
screen "手动设置" 1280x733, template "模板_1"
   on GenerateScreen: SetTag("变量_100", 8)
   Button "HmiScreenItemData_1" at 1116,125 size 159x47; TextOn '向后 / 後向き / 뒤로'; TextOff '向后 / 後向き / 뒤로'
      on Release: ActivateScreen("手动画面", 0)
   IOField "IO 域_20" at 80,185 size 120x41; FormatPattern 99999999
      on Activate: function_f41c6f6c("变量_1")
      ProcessValue <- "ST_HMI_Var_HMI_r64Velocity_Jog_Chuche"
   TextField "文本域_19" at 848,56 size 245x25; Text '当前登录用户 / 目前ログオン中のユーザー / 현재 로그인 사용자'
   IOField "IO 域_15" at 914,98 size 122x41; FormatPattern ?????????????
      ProcessValue <- "user_name"
   IOField "IO 域_2" at 80,417 size 120x41; FormatPattern 99999999
      ProcessValue <- "ST_HMI_Var_HMI_r64Velocity_Jog_JinChe"
   IOField "IO 域_3" at 232,417 size 120x41; FormatPattern 999999999
      ProcessValue <- "ST_HMI_Var_HMI_r64Velocity_Jog_JiaNian"
   IOField "IO 域_5" at 384,417 size 120x41; FormatPattern 999999999
      ProcessValue <- "ST_HMI_Var_HMI_r64Velocity_Jog_JuanRao"
   IOField "IO 域_4" at 232,185 size 120x41; FormatPattern 99999999
      ProcessValue <- "ST_HMI_Var_HMI_r64Velocity_Jog_SongTiao"
   IOField "IO 域_16" at 384,185 size 120x41; FormatPattern 999999999
      ProcessValue <- "ST_HMI_Var_HMI_r64Velocity_Jog_TuiRao"
   IOField "IO 域_6" at 536,416 size 120x41; Authorization "User administration"; FormatPattern 99999999
      ProcessValue <- "ST_HMI_Var_HMI_r64Velocity_Jog_ChengXing_Up"
   IOField "IO 域_7" at 536,186 size 120x41; Authorization "User administration"; FormatPattern 99999999
      ProcessValue <- "ST_HMI_Var_HMI_r64Velocity_Jog_ChengXing_Down"
   IOField "IO 域_9" at 688,184 size 120x41; Authorization "User administration"; FormatPattern 99999999
      ProcessValue <- "ST_HMI_Var_HMI_r64Velocity_Jog_ZhangLi_Up"
   IOField "IO 域_10" at 688,416 size 120x41; Authorization "User administration"; FormatPattern 99999999
      ProcessValue <- "ST_HMI_Var_HMI_r64Velocity_Jog_ZhangLi_Down"
   IOField "IO 域_21" at 80,253 size 120x41; FormatPattern 99999999
      on Activate: function_f41c6f6c("变量_1")
      ProcessValue <- "ST_HMI_Var_HMI_r64AccVelocity_Jog_ChuChe"
   IOField "IO 域_8" at 80,485 size 120x41; FormatPattern 99999999
      ProcessValue <- "ST_HMI_Var_HMI_r64AccVelocity_Jog_JinChe"
   Button "OBJECT_119" at 328,588 size 177x68; TextOff '选择市电模式 / EXIT / 買電モードの選択 / 일반전력'; Authorization "Operate_5"
      on Press: SetBit("ST_HMI_Var_HMI_Bo_Feed_On_Off_Select")
      Appearance <- "ST_HMI_Var_HMI_Bo_Feed_On_Off_Select"
   Button "OBJECT_120" at 573,588 size 177x68; TextOff '选择发电模式 / EXIT / 発電モードの選択 / 발전기 전력'; Authorization "Operate_5"
      on Press: ResetBit("ST_HMI_Var_HMI_Bo_Feed_On_Off_Select")
      Appearance <- "ST_HMI_Var_HMI_Bo_Feed_On_Off_Select"
   Button "OBJECT_5" at 80,80 size 120x80; TextOff '出车 / EXIT / 出機 / 외진'
      on Release: ResetBit("ST_HMI_Var_HMI_bo_ChuChe")
      on Press: SetBit("ST_HMI_Var_HMI_bo_ChuChe")
      Appearance <- "ST_HMI_Var_HMI_bo_ChuChe"
   Button "OBJECT_7" at 232,80 size 120x80; TextOff '送条 / EXIT / 篠送り出し / 시누공급'
      on Release: InvertBit("ST_HMI_Var_HMI_bo_SongTiao")
      Appearance <- "ST_HMI_Var_HMI_bo_SongTiao"
   Button "OBJECT_9" at 384,80 size 120x80; TextOff '退绕 EXIT パッキ ングオフ 언와인딩'
      on Release: ResetBit("ST_HMI_Var_HMI_bo_TuiRao")
      on Press: SetBit("ST_HMI_Var_HMI_bo_TuiRao")
      Appearance <- "ST_HMI_Var_HMI_bo_TuiRao"
   Button "OBJECT_12" at 536,80 size 120x80; TextOff '成形弓降 EXIT ワインデ ィング フォ ーラー下降 성형호랑 하강'
      on Release: ResetBit("ST_HMI_Var_HMI_bo_ChengXing_Down")
      on Press: SetBit("ST_HMI_Var_HMI_bo_ChengXing_Down")
      Appearance <- "ST_HMI_Var_HMI_bo_ChengXing_Down"
   Button "OBJECT_13" at 688,80 size 120x80; TextOff '张力弓升 EXIT カウンタ ーフォー ラー上昇 장력호랑 상승'
      on Release: ResetBit("ST_HMI_Var_HMI_bo_ZhangLi_Up")
      on Press: SetBit("ST_HMI_Var_HMI_bo_ZhangLi_Up")
      Appearance <- "ST_HMI_Var_HMI_bo_ZhangLi_Up"
   Button "OBJECT_6" at 81,312 size 120x80; TextOff '进车 / EXIT / 入機 / 내진'
      on Release: ResetBit("ST_HMI_Var_HMI_bo_JinChe")
      on Press: SetBit("ST_HMI_Var_HMI_bo_JinChe")
      Appearance <- "ST_HMI_Var_HMI_bo_JinChe"
   Button "OBJECT_8" at 232,312 size 120x80; TextOff '加捻 / EXIT / 撚掛 / 연사'
      on Release: ResetBit("ST_HMI_Var_HMI_bo_JiaNian")
      on Press: SetBit("ST_HMI_Var_HMI_bo_JiaNian")
      Appearance <- "ST_Main_Var_g_bo_JianNian_Jog_Status"
   Button "OBJECT_10" at 384,312 size 120x80; TextOff '卷绕 / EXIT / 巻取 / 와인딩'
      on Release: ResetBit("ST_HMI_Var_HMI_bo_JuanRao")
      on Press: SetBit("ST_HMI_Var_HMI_bo_JuanRao")
      Appearance <- "ST_HMI_Var_HMI_bo_JuanRao"
   Button "OBJECT_11" at 536,312 size 120x80; TextOff '成形弓升 EXIT ワインデ ィング フォ ーラー上昇 성형호랑 상승'
      on Release: ResetBit("ST_HMI_Var_HMI_bo_ChengXing_Up")
      on Press: SetBit("ST_HMI_Var_HMI_bo_ChengXing_Up")
      Appearance <- "ST_HMI_Var_HMI_bo_ChengXing_Up"
   Button "OBJECT_14" at 688,312 size 120x80; TextOff '张力弓降 EXIT カウンタ ーフォー ラー下降 장력호랑 하강'
      on Release: ResetBit("ST_HMI_Var_HMI_bo_ZhangLi_Down")
      on Press: SetBit("ST_HMI_Var_HMI_bo_ZhangLi_Down")
      Appearance <- "ST_HMI_Var_HMI_bo_ZhangLi_Down"
   Button "OBJECT_1" at 536,482 size 120x80; TextOff '成形弓 抱闸松开 EXIT'
      on Press: InvertBit("ST_HMI_Var_HMI_bo_ChengXing_Holding_Brake_Open")
      Visibility <- "ST_Main_Var_g_i16_Mode_Enabled"
      ObjectEnable <- "ST_Main_Var_g_i16_Disable_Status"
      Appearance <- "ST_HMI_Var_HMI_bo_ChengXing_Holding_Brake_Open"
   Button "OBJECT_2" at 688,482 size 120x80; TextOff '张力弓 抱闸松开 EXIT'
      on Press: InvertBit("ST_HMI_Var_HMI_bo_ZhangLi_Holding_Brake_Open")
      Visibility <- "ST_Main_Var_g_i16_Mode_Enabled"
      ObjectEnable <- "ST_Main_Var_g_i16_Disable_Status"
      Appearance <- "ST_HMI_Var_HMI_bo_ZhangLi_Holding_Brake_Open"
   Button "OBJECT_3" at 376,481 size 120x80; TextOff '走车 抱闸松开 EXIT'
      on Press: InvertBit("ST_HMI_Var_HMI_bo_ZouChe_Holding_Brake_Open")
      Visibility <- "ST_Main_Var_g_i16_Mode_Enabled"
      ObjectEnable <- "ST_Main_Var_g_i16_Disable_Status"
      Appearance <- "ST_HMI_Var_HMI_bo_ZouChe_Holding_Brake_Open"

screen "牵伸相关" 1280x733, template "模板_3"
   on GenerateScreen: SetTag("变量_100", 15)
   Button "HmiScreenItemData_1" at 1120,10 size 159x47; TextOn '向后 / 뒤로'; TextOff '向后 / 뒤로'
      on Release: ActivateScreen("牵伸调整画面", 0); SetTag("ST_HMI_Var_HMI_i32_ZouChe_ZhanJu_ss_1", 0)
   IOField "IO 域_5" at 346,121 size 126x56; FormatPattern 9.999
      ProcessValue <- "ST_Cam5_Data_Var_g_tz3"
   IOField "IO 域_10" at 61,388 size 114x56; FormatPattern 9.9999
      ProcessValue <- "ST_Cam5_Data_Var_fi"
   IOField "IO 域_11" at 61,317 size 126x55; FormatPattern s9.99
      ProcessValue <- "ST_Cam5_Data_Var_g_ratioV"
   IOField "IO 域_12" at 201,317 size 126x55; FormatPattern 9.99
      ProcessValue <- "ST_Cam5_Data_Var_g_ratioT"
   TextField "文本域_13" at 75,275 size 132x37; Text 'ratioV'
   TextField "文本域_14" at 215,275 size 132x37; Text 'ratioT'
   IOField "IO 域_14" at 343,317 size 126x55; FormatPattern 9.99
      ProcessValue <- "ST_Cam5_Data_Var_g_ratio"
   TextField "文本域_16" at 346,275 size 116x37; Text 'ratio'
   IOField "IO 域_7" at 66,121 size 126x56; FormatPattern 9999
      ProcessValue <- "ST_HMI_Var_HMI_r64Position_ChuChe"
   IOField "IO 域_9" at 66,205 size 126x56; FormatPattern 9.99
      ProcessValue <- "ST_HMI_Var_HMI_r64QianShen_All"
   IOField "IO 域_13" at 206,205 size 126x56; FormatPattern 9.99
      ProcessValue <- "ST_HMI_Var_HMI_r64QianShen_First"
   IOField "IO 域_15" at 346,205 size 126x56; FormatPattern 999
      ProcessValue <- "ST_HMI_Var_HMI_r64QianShen_FirstArea"
   IOField "IO 域_16" at 486,205 size 126x56; FormatPattern 99
      ProcessValue <- "ST_HMI_Var_HMI_r64QianShen_finalArea"
   Button "Button" at 500,121 size 98x56; TextOff 'CAM5'
      Appearance <- "Cam_5_accessState"
   IOField "IO 域_8" at 206,121 size 126x56; FormatPattern 999
      ProcessValue <- "ST_Cam5_Data_Var_g_vm"
   IOField "IO 域_1" at 1104,96 size 126x56; FormatPattern 9999999999
      ProcessValue <- "ST_HMI_Var_HMI_i32_ZouChe_ZhanJu_ss_1"
   IOField "IO 域_2" at 1104,168 size 126x56; FormatPattern 9999
      ProcessValue <- "ST_HMI_Var_HMI_r64_ZouChe_ZhanJu_Max_20"
      Visibility <- "ST_HMI_Var_HMI_bo_ZouChe_ZhanJu_Select"
   IOField "IO 域_3" at 1104,240 size 126x56; FormatPattern 9999
      ProcessValue <- "ST_HMI_Var_HMI_r64_ZouChe_ZhanJu_Max_25"
      Visibility <- "ST_HMI_Var_HMI_bo_ZouChe_ZhanJu_Select"
   IOField "IO 域_4" at 1104,312 size 126x56; FormatPattern 9999
      ProcessValue <- "ST_HMI_Var_HMI_r64_ZouChe_ZhanJu_Max_30"
      Visibility <- "ST_HMI_Var_HMI_bo_ZouChe_ZhanJu_Select"
   IOField "IO 域_6" at 1104,384 size 126x56; FormatPattern 9999
      ProcessValue <- "ST_HMI_Var_HMI_r64_ZouChe_ZhanJu_Max_35"
      Visibility <- "ST_HMI_Var_HMI_bo_ZouChe_ZhanJu_Select"
   IOField "IO 域_17" at 1104,456 size 126x56; FormatPattern 9999
      ProcessValue <- "ST_HMI_Var_HMI_r64_ZouChe_ZhanJu_Max_40"
      Visibility <- "ST_HMI_Var_HMI_bo_ZouChe_ZhanJu_Select"
   IOField "IO 域_18" at 1104,528 size 126x56; FormatPattern 9999
      ProcessValue <- "ST_HMI_Var_HMI_r64_ZouChe_ZhanJu_Max_45"
      Visibility <- "ST_HMI_Var_HMI_bo_ZouChe_ZhanJu_Select"
   IOField "IO 域_19" at 1104,600 size 126x56; FormatPattern 9999
      ProcessValue <- "ST_HMI_Var_HMI_r64_ZouChe_ZhanJu_Max_Effect"
      Visibility <- "ST_HMI_Var_HMI_bo_ZouChe_ZhanJu_Select"
   Button "Button_1" at 960,168 size 126x56; TextOff '2.0米'
      on Release: SetTag("ST_HMI_Var_HMI_i16_ZouChe_ZhanJu_Select", 20)
      Appearance <- "ST_HMI_Var_HMI_i16_ZouChe_ZhanJu_Select"
      Visibility <- "ST_HMI_Var_HMI_bo_ZouChe_ZhanJu_Select"
   Button "Button_2" at 960,240 size 126x56; TextOff '2.5米'
      on Release: SetTag("ST_HMI_Var_HMI_i16_ZouChe_ZhanJu_Select", 25)
      Appearance <- "ST_HMI_Var_HMI_i16_ZouChe_ZhanJu_Select"
      Visibility <- "ST_HMI_Var_HMI_bo_ZouChe_ZhanJu_Select"
   Button "Button_3" at 960,312 size 126x56; TextOff '3.0米'
      on Release: SetTag("ST_HMI_Var_HMI_i16_ZouChe_ZhanJu_Select", 30)
      Appearance <- "ST_HMI_Var_HMI_i16_ZouChe_ZhanJu_Select"
      Visibility <- "ST_HMI_Var_HMI_bo_ZouChe_ZhanJu_Select"
   Button "Button_4" at 960,384 size 126x56; TextOff '3.5米'
      on Release: SetTag("ST_HMI_Var_HMI_i16_ZouChe_ZhanJu_Select", 35)
      Appearance <- "ST_HMI_Var_HMI_i16_ZouChe_ZhanJu_Select"
      Visibility <- "ST_HMI_Var_HMI_bo_ZouChe_ZhanJu_Select"
   Button "Button_5" at 960,456 size 126x56; TextOff '4.0米'
      on Release: SetTag("ST_HMI_Var_HMI_i16_ZouChe_ZhanJu_Select", 40)
      Appearance <- "ST_HMI_Var_HMI_i16_ZouChe_ZhanJu_Select"
      Visibility <- "ST_HMI_Var_HMI_bo_ZouChe_ZhanJu_Select"
   Button "Button_6" at 960,528 size 126x56; TextOff '4.5米'
      on Release: SetTag("ST_HMI_Var_HMI_i16_ZouChe_ZhanJu_Select", 45)
      Appearance <- "ST_HMI_Var_HMI_i16_ZouChe_ZhanJu_Select"
      Visibility <- "ST_HMI_Var_HMI_bo_ZouChe_ZhanJu_Select"
   Button "Button_7" at 960,600 size 126x56; TextOff '生效'
      Visibility <- "ST_HMI_Var_HMI_bo_ZouChe_ZhanJu_Select"

Template "Template_1" 1280x733
   Button "Template_Button_1" at 1200,64 size 78x59; TextOn 'Login'; TextOff 'Login'; PictureOn "Login_TP1200_Comfort"; PictureOff "Login_TP1200_Comfort"
      on Release: function_a2a04561()
   Button "Template_Button_2" at 1200,126 size 78x59; TextOn 'AlarmDisplay'; TextOff 'AlarmDisplay'; PictureOn "AlarmDisplay_TP1200_Comfort"; PictureOff "AlarmDisplay_TP1200_Comfort"
   Button "Template_Button_3" at 1200,187 size 78x59; TextOn 'ToggleLanguage'; TextOff 'ToggleLanguage'; PictureOn "ToggleLanguage_TP1200_Comfort"; PictureOff "ToggleLanguage_TP1200_Comfort"
      on Release: function_fb9197e8(-1)
   Button "Template_Button_4" at 1200,249 size 78x59; TextOff 'Text'
   Button "Template_Button_5" at 1200,310 size 78x59; TextOff 'Text'
   Button "Template_Button_6" at 1200,372 size 78x59; TextOff 'Text'
   Button "Template_Button_7" at 1200,433 size 78x59; TextOff 'Text'
   Button "Template_Button_8" at 1200,495 size 78x59; TextOff 'Text'
   Button "Template_Button_9" at 1200,556 size 78x59; TextOff 'Text'
   Button "Template_Button_10" at 1200,618 size 78x59; TextOff 'Text'
   Button "Template_Button_11" at 1200,679 size 78x59; TextOn 'NavigateHome'; TextOff 'NavigateHome'; PictureOn "NavigateHome_TP1200_Comfort"; PictureOff "NavigateHome_TP1200_Comfort"
      on Release: ActivateScreen("自动画面", 0)
   Button "Template_Button_12" at 1200,2 size 78x59; TextOff 'Text'; PictureOff "1"
      on Click: StopRuntime(0)

Template "模板_2" 1280x733
   Button "Template_Button_11" at 1200,673 size 78x59; TextOn 'NavigateHome'; TextOff 'NavigateHome'; PictureOn "NavigateHome_TP1200_Comfort"; PictureOff "NavigateHome_TP1200_Comfort"
      on Release: ActivateScreen("自动画面", 0)
      on Press: function_f23ef4c9()

Template "模板_1" 1280x733
   Button "Template_Button_11" at 1200,673 size 78x59; TextOn 'NavigateHome'; TextOff 'NavigateHome'; PictureOn "NavigateHome_TP1200_Comfort"; PictureOff "NavigateHome_TP1200_Comfort"
      on Release: ActivateScreen("自动画面", 0); SetTag("ST_HMI_Var_HMI_i32_ZouChe_ZhanJu_ss_1", 0)
      on Press: function_f23ef4c9()

Template "模板_3" 1280x733
   Button "Template_Button_11" at 1200,673 size 78x59; TextOn 'NavigateHome'; TextOff 'NavigateHome'; PictureOn "NavigateHome_TP1200_Comfort"; PictureOff "NavigateHome_TP1200_Comfort"
      on Release: ActivateScreen("自动画面", 0); SetTag("ST_HMI_Var_HMI_i32_ZouChe_ZhanJu_ss_1", 0)
      on Press: function_f23ef4c9()

screen "纱穗参数设定" 1280x733, template "模板_2"
   Button "HmiScreenItemData_1" at 1121,79 size 159x47; TextOn '向后 / 뒤로'; TextOff '向后 / 뒤로'
      on Release: ActivateScreen("常用调试画面", 0); function_f23ef4c9()
   TextField "Text Field_50" at 136,234 size 384x56; Text '总高度H: / 총높이H'
   TextField "Text Field_51" at 136,304 size 384x56; Text '上锥体高度HS2: / 상단 코프높이HS2'
   TextField "Text Field_52" at 311,24 size 280x42; Text '纱穗参数设定 / 코프 형성'
   TextField "Text Field_53" at 136,374 size 384x56; Text '上锥体高度HS2_D: / 상단 코프높이M (중간)HS2_D'
   TextField "Text Field_55" at 732,162 size 67x56; Text 'mm'
   TextField "Text Field_56" at 732,232 size 67x56; Text 'mm'
   TextField "Text Field_57" at 732,302 size 67x56; Text 'mm'
   TextField "Text Field_58" at 732,372 size 67x56; Text 'mm'
   TextField "Text Field_59" at 136,444 size 384x56; Text '最大直径D: / 최대 직경D'
   TextField "Text Field_60" at 732,442 size 67x56; Text 'mm'
   TextField "Text Field_54" at 136,94 size 384x56; Text '起始点高度Hqs: / 출발점 높이Hqs'
   TextField "Text Field_61" at 732,92 size 67x56; Text 'mm'
   TextField "Text Field_62" at 136,164 size 384x56; Text '下锥体高度Hs1: / 하부높이HS1'
   IOField "IO Field_27" at 550,232 size 140x56; FormatPattern 999.9
      ProcessValue <- "ST_HMI_Var_HMI_r64Height_ShaSui_whole"
   IOField "IO Field_28" at 550,302 size 140x56; FormatPattern 99.9
      ProcessValue <- "ST_HMI_Var_HMI_r64Height_ShaSui_Top"
   IOField "IO Field_29" at 550,372 size 140x56; FormatPattern 99.9
      ProcessValue <- "ST_HMI_Var_HMI_r64Height_ShaSui_Top_MaxD"
   IOField "IO Field_30" at 550,442 size 140x56; FormatPattern 99.9
      ProcessValue <- "ST_HMI_Var_HMI_r64Diameter_ShaSui_Max"
   IOField "IO Field_31" at 550,92 size 140x56; FormatPattern 99.9
      ProcessValue <- "ST_HMI_Var_HMI_r64Height_ShaSui_Start"
   IOField "IO Field_32" at 550,162 size 140x56; FormatPattern 99.9
      ProcessValue <- "ST_HMI_Var_HMI_r64Height_ShaSui_Bottom"

screen "监控画面" 1280x733, template "模板_2"
   IOField "IO Field_3" at 48,24 size 128x42; FormatPattern 99.999
      ProcessValue <- "ST_Real_Monitoring_HMI_r64_Real_QianShen_WuNian"
   IOField "IO Field_1" at 48,80 size 128x42; FormatPattern 99.999
      ProcessValue <- "ST_HMI_Var_HMI_r64QianShen_All_real"
   IOField "IO Field_2" at 48,144 size 128x42; FormatPattern 9999.99
      ProcessValue <- "ST_Real_Monitoring_HMI_r64Axis_ZouChe_Position_JiZhong_QianShen_Start"
   IOField "IO Field_4" at 48,200 size 128x42; FormatPattern 9999
      ProcessValue <- "ST_Real_Monitoring_HMI_r64_NianDu_JiZhong_QianShen_Start"
   IOField "IO Field_5" at 48,264 size 128x42; FormatPattern 9999.99
      ProcessValue <- "ST_Real_Monitoring_HMI_r64Axis_ZouChe_Position_LuoLa_Stop"
   IOField "IO Field_6" at 48,320 size 128x42; FormatPattern 9999
      ProcessValue <- "ST_Real_Monitoring_HMI_r64_NianDu_LuoLa_Stop"
   IOField "IO Field_7" at 48,384 size 128x42; FormatPattern 9999
      ProcessValue <- "ST_HMI_Var_HMI_r64NianDu_actual"
   IOField "IO Field_8" at 48,440 size 128x42; FormatPattern 9999.99
      ProcessValue <- "ST_Real_Monitoring_HMI_r64Axis_ZouChe_Position_YiNian_DaoDa"
   Button "HmiScreenItemData_1" at 1106,176 size 145x54; TextOn '向后 / 後向き / 뒤로'; TextOff '向后 / 後向き / 뒤로'
      on Release: ActivateScreen("设置画面", 0); function_f23ef4c9()
   IOField "IO Field_10" at 588,24 size 128x42; FormatPattern 99.999
      ProcessValue <- "ST_Convert_ReadParameters_g_r64_SERVO_03_ZouChe_35_Motor_temperature_real"
   IOField "IO Field_11" at 588,82 size 128x42; FormatPattern 999.99
      ProcessValue <- "ST_Convert_ReadParameters_g_r64_SERVO_04_ZhangLi_35_Motor_temperature_real"
   IOField "IO Field_12" at 588,144 size 128x42; FormatPattern 999.99
      ProcessValue <- "ST_Convert_ReadParameters_g_r64_SERVO_05_ChengXing_35_Motor_temperature_real"
   IOField "IO Field_13" at 588,200 size 128x42; FormatPattern 999.99
      ProcessValue <- "ST_Convert_ReadParameters_g_r64_SERVO_06_GunTong_35_Motor_temperature_real"
   IOField "IO Field_14" at 588,264 size 128x42; FormatPattern 999.99
      ProcessValue <- "ST_Convert_ReadParameters_g_r64_SERVO_08_LuoLa_35_Motor_temperature_real"
   IOField "IO Field_15" at 588,320 size 128x42; FormatPattern 999.99
      ProcessValue <- "ST_Convert_ReadParameters_g_r64_SERVO_07_DingZi_35_Motor_temperature_real"
   IOField "IO Field_17" at 588,370 size 128x42; FormatPattern 999.99
      ProcessValue <- "ST_Convert_ReadParameters_g_r64_SERVO_03_ZouChe_37_4_Power_unit_temperatures_Interior_of_power_unit_real"
   IOField "IO Field_18" at 588,426 size 128x42; FormatPattern 999.99
      ProcessValue <- "ST_Convert_ReadParameters_g_r64_SERVO_05_ChengXing_37_4_Power_unit_temperatures_Interior_of_power_unit_real"
   IOField "IO Field_19" at 588,482 size 128x42; FormatPattern 999.99
      ProcessValue <- "ST_Convert_ReadParameters_g_r64_SERVO_07_DingZi_37_4_Power_unit_temperatures_Interior_of_power_unit_real"
   IOField "IO Field_20" at 588,538 size 128x42; FormatPattern 999.99
      ProcessValue <- "ST_Convert_ReadParameters_g_r64_SERVO_08_LuoLa_37_4_Power_unit_temperatures_Interior_of_power_unit_real"
   TextField "Text Field_40" at 191,24 size 352x42; Text '实时无捻牵伸 / 番手: / 실 번수'
   TextField "Text Field_1" at 193,80 size 352x42; Text '实时总牵伸 / 番手: / 실 번수'
   TextField "Text Field_2" at 194,144 size 352x42; Text '集中牵伸开始时的走车位置 / 番手: / 실 번수'
   TextField "Text Field_3" at 193,200 size 352x42; Text '集中牵伸开始时的捻度 / 番手: / 실 번수'
   TextField "Text Field_4" at 195,264 size 352x42; Text '罗拉停止时的走车位置 / 番手: / 실 번수'
   TextField "Text Field_5" at 194,320 size 352x42; Text '罗拉停止时的捻度 / 番手: / 실 번수'
   TextField "Text Field_6" at 194,384 size 352x42; Text '实际捻度 / 番手: / 실 번수'
   TextField "Text Field_7" at 193,440 size 352x42; Text '锭子加速到第一个峰值时的走车位置 / 番手: / 실 번수'
   TextField "Text Field_9" at 732,24 size 352x42; Text '走车电机实时温度（℃） / 番手: / 실 번수'
   TextField "Text Field_10" at 732,82 size 352x42; Text '张力电机实时温度（℃） / 番手: / 실 번수'
   TextField "Text Field_11" at 732,144 size 352x42; Text '成形电机实时温度（℃） / 番手: / 실 번수'
   TextField "Text Field_12" at 732,200 size 352x42; Text '滚筒电机实时温度（℃） / 番手: / 실 번수'
   TextField "Text Field_13" at 732,264 size 352x42; Text '罗拉电机实时温度（℃） / 番手: / 실 번수'
   TextField "Text Field_14" at 732,320 size 352x42; Text '锭子电机实时温度（℃） / 番手: / 실 번수'
   TextField "Text Field_16" at 732,370 size 352x42; Text '走车张力驱动器实时温度（℃） / 番手: / 실 번수'
   TextField "Text Field_17" at 732,426 size 352x42; Text '成形滚筒驱动器实时温度（℃） / 番手: / 실 번수'
   TextField "Text Field_18" at 732,482 size 352x42; Text '锭子驱动器实时温度（℃） / 番手: / 실 번수'
   TextField "Text Field_19" at 732,538 size 352x42; Text '罗拉驱动器实时温度（℃） / 番手: / 실 번수'

screen "用户管理" 1280x733, template "模板_2"
   on GenerateScreen: SetTag("变量_100", 21)
   Button "HmiScreenItemData_1" at 1119,57 size 159x47; TextOn '向后'; TextOff '向后'
      on Release: ActivateScreen("自动画面", 0); function_f23ef4c9()
   Button "Button_1" at 890,57 size 170x60; TextOff '登录用户'
      on Press: function_a2a04561()
   Button "Button_2" at 890,181 size 170x60; TextOff '注销用户'
      on Press: function_f23ef4c9()
   UserView "用户视图_1" at 2,1 size 858x730
   UserView "HmiScreenItemData" at 1,0 size 862x729

screen "卷绕经验参数" 1280x733, template "模板_2"
   on GenerateScreen: SetTag("变量_100", 20)
   IOField "IO Field_41" at 24,65 size 112x38; FormatPattern 99.99
      ProcessValue <- "ST_Calculation_Var_1_ZhiShu_ARRAY_JR{3}"
   IOField "IO Field_1" at 156,64 size 112x38; FormatPattern 99.999
      ProcessValue <- "ST_Calculation_Var_1_f1_n_delt_0_n_ARRAY_JR{3}"
   IOField "IO Field_2" at 288,64 size 112x38; FormatPattern 99.999
      ProcessValue <- "ST_Calculation_Var_1_g1_n_delt_0_n_ARRAY_JR{3}"
   IOField "IO Field_3" at 24,108 size 112x38; FormatPattern 99.99
      ProcessValue <- "ST_Calculation_Var_1_ZhiShu_ARRAY_JR{4}"
   IOField "IO Field_4" at 156,108 size 112x38; FormatPattern 99.999
      ProcessValue <- "ST_Calculation_Var_1_f1_n_delt_0_n_ARRAY_JR{4}"
   IOField "IO Field_5" at 288,108 size 112x38; FormatPattern 99.999
      ProcessValue <- "ST_Calculation_Var_1_g1_n_delt_0_n_ARRAY_JR{4}"
   IOField "IO Field_6" at 24,153 size 112x38; FormatPattern 99.99
      ProcessValue <- "ST_Calculation_Var_1_ZhiShu_ARRAY_JR{5}"
   IOField "IO Field_7" at 24,197 size 112x38; FormatPattern 99.99
      ProcessValue <- "ST_Calculation_Var_1_ZhiShu_ARRAY_JR{6}"
   IOField "IO Field_8" at 24,242 size 112x38; FormatPattern 99.99
      ProcessValue <- "ST_Calculation_Var_1_ZhiShu_ARRAY_JR{7}"
   IOField "IO Field_9" at 24,286 size 112x38; FormatPattern 99.99
      ProcessValue <- "ST_Calculation_Var_1_ZhiShu_ARRAY_JR{8}"
   IOField "IO Field_10" at 24,331 size 112x38; FormatPattern 99.99
      ProcessValue <- "ST_Calculation_Var_1_ZhiShu_ARRAY_JR{9}"
   IOField "IO Field_11" at 24,376 size 112x38; FormatPattern 99.99
      ProcessValue <- "ST_Calculation_Var_1_ZhiShu_ARRAY_JR{10}"
   IOField "IO Field_12" at 24,420 size 112x38; FormatPattern 99.99
      ProcessValue <- "ST_Calculation_Var_1_ZhiShu_ARRAY_JR{11}"
   IOField "IO Field_13" at 24,465 size 112x38; FormatPattern 99.99
      ProcessValue <- "ST_Calculation_Var_1_ZhiShu_ARRAY_JR{12}"
   IOField "IO Field_14" at 24,509 size 112x38; FormatPattern 99.99
      ProcessValue <- "ST_Calculation_Var_1_ZhiShu_ARRAY_JR{13}"
   IOField "IO Field_15" at 24,554 size 112x38; FormatPattern 99.99
      ProcessValue <- "ST_Calculation_Var_1_ZhiShu_ARRAY_JR{14}"
   IOField "IO Field_16" at 24,598 size 112x38; FormatPattern 99.99
      ProcessValue <- "ST_Calculation_Var_1_ZhiShu_ARRAY_JR{15}"
   IOField "IO Field_17" at 24,643 size 112x38; FormatPattern 99.99
      ProcessValue <- "ST_Calculation_Var_1_ZhiShu_ARRAY_JR{16}"
   IOField "IO Field_18" at 24,688 size 112x38; FormatPattern 99.99
      ProcessValue <- "ST_Calculation_Var_1_ZhiShu_ARRAY_JR{17}"
   IOField "IO Field_19" at 156,153 size 112x38; FormatPattern 99.999
      ProcessValue <- "ST_Calculation_Var_1_f1_n_delt_0_n_ARRAY_JR{5}"
   IOField "IO Field_20" at 156,197 size 112x38; FormatPattern 99.999
      ProcessValue <- "ST_Calculation_Var_1_f1_n_delt_0_n_ARRAY_JR{6}"
   IOField "IO Field_21" at 156,242 size 112x38; FormatPattern 99.999
      ProcessValue <- "ST_Calculation_Var_1_f1_n_delt_0_n_ARRAY_JR{7}"
   IOField "IO Field_22" at 156,286 size 112x38; FormatPattern 99.999
      ProcessValue <- "ST_Calculation_Var_1_f1_n_delt_0_n_ARRAY_JR{8}"
   IOField "IO Field_23" at 156,331 size 112x38; FormatPattern 99.999
      ProcessValue <- "ST_Calculation_Var_1_f1_n_delt_0_n_ARRAY_JR{9}"
   IOField "IO Field_24" at 156,376 size 112x38; FormatPattern 99.999
      ProcessValue <- "ST_Calculation_Var_1_f1_n_delt_0_n_ARRAY_JR{10}"
   IOField "IO Field_25" at 156,420 size 112x38; FormatPattern 99.999
      ProcessValue <- "ST_Calculation_Var_1_f1_n_delt_0_n_ARRAY_JR{11}"
   IOField "IO Field_26" at 156,465 size 112x38; FormatPattern 99.999
      ProcessValue <- "ST_Calculation_Var_1_f1_n_delt_0_n_ARRAY_JR{12}"
   IOField "IO Field_27" at 156,509 size 112x38; FormatPattern 99.999
      ProcessValue <- "ST_Calculation_Var_1_f1_n_delt_0_n_ARRAY_JR{13}"
   IOField "IO Field_28" at 156,554 size 112x38; FormatPattern 99.999
      ProcessValue <- "ST_Calculation_Var_1_f1_n_delt_0_n_ARRAY_JR{14}"
   IOField "IO Field_29" at 156,598 size 112x38; FormatPattern 99.999
      ProcessValue <- "ST_Calculation_Var_1_f1_n_delt_0_n_ARRAY_JR{15}"
   IOField "IO Field_30" at 156,643 size 112x38; FormatPattern 99.999
      ProcessValue <- "ST_Calculation_Var_1_f1_n_delt_0_n_ARRAY_JR{16}"
   IOField "IO Field_31" at 156,688 size 112x38; FormatPattern 99.999
      ProcessValue <- "ST_Calculation_Var_1_f1_n_delt_0_n_ARRAY_JR{17}"
   IOField "IO Field_32" at 288,153 size 112x38; FormatPattern 99.999
      ProcessValue <- "ST_Calculation_Var_1_g1_n_delt_0_n_ARRAY_JR{5}"
   IOField "IO Field_33" at 288,197 size 112x38; FormatPattern 99.999
      ProcessValue <- "ST_Calculation_Var_1_g1_n_delt_0_n_ARRAY_JR{6}"
   IOField "IO Field_34" at 288,242 size 112x38; FormatPattern 99.999
      ProcessValue <- "ST_Calculation_Var_1_g1_n_delt_0_n_ARRAY_JR{7}"
   IOField "IO Field_35" at 288,286 size 112x38; FormatPattern 99.999
      ProcessValue <- "ST_Calculation_Var_1_g1_n_delt_0_n_ARRAY_JR{8}"
   IOField "IO Field_36" at 288,331 size 112x38; FormatPattern 99.999
      ProcessValue <- "ST_Calculation_Var_1_g1_n_delt_0_n_ARRAY_JR{9}"
   IOField "IO Field_37" at 288,376 size 112x38; FormatPattern 99.999
      ProcessValue <- "ST_Calculation_Var_1_g1_n_delt_0_n_ARRAY_JR{10}"
   IOField "IO Field_38" at 288,420 size 112x38; FormatPattern 99.999
      ProcessValue <- "ST_Calculation_Var_1_g1_n_delt_0_n_ARRAY_JR{11}"
   IOField "IO Field_39" at 288,465 size 112x38; FormatPattern 99.999
      ProcessValue <- "ST_Calculation_Var_1_g1_n_delt_0_n_ARRAY_JR{12}"
   IOField "IO Field_40" at 288,509 size 112x38; FormatPattern 99.999
      ProcessValue <- "ST_Calculation_Var_1_g1_n_delt_0_n_ARRAY_JR{13}"
   IOField "IO Field_42" at 288,554 size 112x38; FormatPattern 99.999
      ProcessValue <- "ST_Calculation_Var_1_g1_n_delt_0_n_ARRAY_JR{14}"
   IOField "IO Field_43" at 288,598 size 112x38; FormatPattern 99.999
      ProcessValue <- "ST_Calculation_Var_1_g1_n_delt_0_n_ARRAY_JR{15}"
   IOField "IO Field_44" at 288,643 size 112x38; FormatPattern 99.999
      ProcessValue <- "ST_Calculation_Var_1_g1_n_delt_0_n_ARRAY_JR{16}"
   IOField "IO Field_45" at 288,688 size 112x38; FormatPattern 99.999
      ProcessValue <- "ST_Calculation_Var_1_g1_n_delt_0_n_ARRAY_JR{17}"
   IOField "IO Field_46" at 420,65 size 112x38; FormatPattern 99.99
      ProcessValue <- "ST_Calculation_Var_1_ZhiShu_ARRAY_JR{18}"
   IOField "IO Field_47" at 552,64 size 112x38; FormatPattern 99.999
      ProcessValue <- "ST_Calculation_Var_1_f1_n_delt_0_n_ARRAY_JR{18}"
   IOField "IO Field_48" at 684,64 size 112x38; FormatPattern 99.999
      ProcessValue <- "ST_Calculation_Var_1_g1_n_delt_0_n_ARRAY_JR{18}"
   IOField "IO Field_49" at 420,108 size 112x38; FormatPattern 99.99
      ProcessValue <- "ST_Calculation_Var_1_ZhiShu_ARRAY_JR{19}"
   IOField "IO Field_50" at 552,108 size 112x38; FormatPattern 99.999
      ProcessValue <- "ST_Calculation_Var_1_f1_n_delt_0_n_ARRAY_JR{19}"
   IOField "IO Field_51" at 684,108 size 112x38; FormatPattern 99.999
      ProcessValue <- "ST_Calculation_Var_1_g1_n_delt_0_n_ARRAY_JR{19}"
   IOField "IO Field_52" at 420,153 size 112x38; FormatPattern 99.99
      ProcessValue <- "ST_Calculation_Var_1_ZhiShu_ARRAY_JR{20}"
   IOField "IO Field_53" at 420,197 size 112x38; FormatPattern 99.99
      ProcessValue <- "ST_Calculation_Var_1_ZhiShu_ARRAY_JR{21}"
   IOField "IO Field_54" at 420,242 size 112x38; FormatPattern 99.99
      ProcessValue <- "ST_Calculation_Var_1_ZhiShu_ARRAY_JR{22}"
   IOField "IO Field_55" at 420,286 size 112x38; FormatPattern 99.99
      ProcessValue <- "ST_Calculation_Var_1_ZhiShu_ARRAY_JR{23}"
   IOField "IO Field_56" at 420,331 size 112x38; FormatPattern 99.99
      ProcessValue <- "ST_Calculation_Var_1_ZhiShu_ARRAY_JR{24}"
   IOField "IO Field_57" at 420,376 size 112x38; FormatPattern 99.99
      ProcessValue <- "ST_Calculation_Var_1_ZhiShu_ARRAY_JR{25}"
   IOField "IO Field_58" at 420,420 size 112x38; FormatPattern 99.99
      ProcessValue <- "ST_Calculation_Var_1_ZhiShu_ARRAY_JR{26}"
   IOField "IO Field_59" at 420,465 size 112x38; FormatPattern 99.99
      ProcessValue <- "ST_Calculation_Var_1_ZhiShu_ARRAY_JR{27}"
   IOField "IO Field_60" at 420,509 size 112x38; FormatPattern 99.99
      ProcessValue <- "ST_Calculation_Var_1_ZhiShu_ARRAY_JR{28}"
   IOField "IO Field_61" at 420,554 size 112x38; FormatPattern 99.99
      ProcessValue <- "ST_Calculation_Var_1_ZhiShu_ARRAY_JR{29}"
   IOField "IO Field_62" at 420,598 size 112x38; FormatPattern 99.99
      ProcessValue <- "ST_Calculation_Var_1_ZhiShu_ARRAY_JR{30}"
   IOField "IO Field_63" at 420,643 size 112x38; FormatPattern 99.99
      ProcessValue <- "ST_Calculation_Var_1_ZhiShu_ARRAY_JR{31}"
   IOField "IO Field_64" at 420,688 size 112x38; FormatPattern 99.99
      ProcessValue <- "ST_Calculation_Var_1_ZhiShu_ARRAY_JR{32}"
   IOField "IO Field_65" at 552,153 size 112x38; FormatPattern 99.999
      ProcessValue <- "ST_Calculation_Var_1_f1_n_delt_0_n_ARRAY_JR{20}"
   IOField "IO Field_66" at 552,197 size 112x38; FormatPattern 99.999
      ProcessValue <- "ST_Calculation_Var_1_f1_n_delt_0_n_ARRAY_JR{21}"
   IOField "IO Field_67" at 552,242 size 112x38; FormatPattern 99.999
      ProcessValue <- "ST_Calculation_Var_1_f1_n_delt_0_n_ARRAY_JR{22}"
   IOField "IO Field_68" at 552,286 size 112x38; FormatPattern 99.999
      ProcessValue <- "ST_Calculation_Var_1_f1_n_delt_0_n_ARRAY_JR{23}"
   IOField "IO Field_69" at 552,331 size 112x38; FormatPattern 99.999
      ProcessValue <- "ST_Calculation_Var_1_f1_n_delt_0_n_ARRAY_JR{24}"
   IOField "IO Field_70" at 552,376 size 112x38; FormatPattern 99.999
      ProcessValue <- "ST_Calculation_Var_1_f1_n_delt_0_n_ARRAY_JR{25}"
   IOField "IO Field_71" at 552,420 size 112x38; FormatPattern 99.999
      ProcessValue <- "ST_Calculation_Var_1_f1_n_delt_0_n_ARRAY_JR{26}"
   IOField "IO Field_72" at 552,465 size 112x38; FormatPattern 99.999
      ProcessValue <- "ST_Calculation_Var_1_f1_n_delt_0_n_ARRAY_JR{27}"
   IOField "IO Field_73" at 552,509 size 112x38; FormatPattern 99.999
      ProcessValue <- "ST_Calculation_Var_1_f1_n_delt_0_n_ARRAY_JR{28}"
   IOField "IO Field_74" at 552,554 size 112x38; FormatPattern 99.999
      ProcessValue <- "ST_Calculation_Var_1_f1_n_delt_0_n_ARRAY_JR{29}"
   IOField "IO Field_75" at 552,598 size 112x38; FormatPattern 99.999
      ProcessValue <- "ST_Calculation_Var_1_f1_n_delt_0_n_ARRAY_JR{30}"
   IOField "IO Field_76" at 552,643 size 112x38; FormatPattern 99.999
      ProcessValue <- "ST_Calculation_Var_1_f1_n_delt_0_n_ARRAY_JR{31}"
   IOField "IO Field_77" at 552,688 size 112x38; FormatPattern 99.999
      ProcessValue <- "ST_Calculation_Var_1_f1_n_delt_0_n_ARRAY_JR{32}"
   IOField "IO Field_78" at 684,153 size 112x38; FormatPattern 99.999
      ProcessValue <- "ST_Calculation_Var_1_g1_n_delt_0_n_ARRAY_JR{20}"
   IOField "IO Field_79" at 684,197 size 112x38; FormatPattern 99.999
      ProcessValue <- "ST_Calculation_Var_1_g1_n_delt_0_n_ARRAY_JR{21}"
   IOField "IO Field_80" at 684,242 size 112x38; FormatPattern 99.999
      ProcessValue <- "ST_Calculation_Var_1_g1_n_delt_0_n_ARRAY_JR{22}"
   IOField "IO Field_81" at 684,286 size 112x38; FormatPattern 99.999
      ProcessValue <- "ST_Calculation_Var_1_g1_n_delt_0_n_ARRAY_JR{23}"
   IOField "IO Field_82" at 684,331 size 112x38; FormatPattern 99.999
      ProcessValue <- "ST_Calculation_Var_1_g1_n_delt_0_n_ARRAY_JR{24}"
   IOField "IO Field_83" at 684,376 size 112x38; FormatPattern 99.999
      ProcessValue <- "ST_Calculation_Var_1_g1_n_delt_0_n_ARRAY_JR{25}"
   IOField "IO Field_84" at 684,420 size 112x38; FormatPattern 99.999
      ProcessValue <- "ST_Calculation_Var_1_g1_n_delt_0_n_ARRAY_JR{26}"
   IOField "IO Field_85" at 684,465 size 112x38; FormatPattern 99.999
      ProcessValue <- "ST_Calculation_Var_1_g1_n_delt_0_n_ARRAY_JR{27}"
   IOField "IO Field_86" at 684,509 size 112x38; FormatPattern 99.999
      ProcessValue <- "ST_Calculation_Var_1_g1_n_delt_0_n_ARRAY_JR{28}"
   IOField "IO Field_87" at 684,554 size 112x38; FormatPattern 99.999
      ProcessValue <- "ST_Calculation_Var_1_g1_n_delt_0_n_ARRAY_JR{29}"
   IOField "IO Field_88" at 684,598 size 112x38; FormatPattern 99.999
      ProcessValue <- "ST_Calculation_Var_1_g1_n_delt_0_n_ARRAY_JR{30}"
   IOField "IO Field_89" at 684,643 size 112x38; FormatPattern 99.999
      ProcessValue <- "ST_Calculation_Var_1_g1_n_delt_0_n_ARRAY_JR{31}"
   IOField "IO Field_90" at 684,688 size 112x38; FormatPattern 99.999
      ProcessValue <- "ST_Calculation_Var_1_g1_n_delt_0_n_ARRAY_JR{32}"
   IOField "IO Field_91" at 816,65 size 112x38; FormatPattern 99.99
      ProcessValue <- "ST_Calculation_Var_1_ZhiShu_ARRAY_JR{33}"
   IOField "IO Field_92" at 948,64 size 112x38; FormatPattern 99.999
      ProcessValue <- "ST_Calculation_Var_1_f1_n_delt_0_n_ARRAY_JR{33}"
   IOField "IO Field_93" at 1080,64 size 112x38; FormatPattern 99.999
      ProcessValue <- "ST_Calculation_Var_1_g1_n_delt_0_n_ARRAY_JR{33}"
   IOField "IO Field_94" at 816,108 size 112x38; FormatPattern 99.99
      ProcessValue <- "ST_Calculation_Var_1_ZhiShu_ARRAY_JR{34}"
   IOField "IO Field_95" at 948,108 size 112x38; FormatPattern 99.999
      ProcessValue <- "ST_Calculation_Var_1_f1_n_delt_0_n_ARRAY_JR{34}"
   IOField "IO Field_96" at 1080,108 size 112x38; FormatPattern 99.999
      ProcessValue <- "ST_Calculation_Var_1_g1_n_delt_0_n_ARRAY_JR{34}"
   IOField "IO Field_97" at 816,153 size 112x38; FormatPattern 99.99
      ProcessValue <- "ST_Calculation_Var_1_ZhiShu_ARRAY_JR{35}"
   IOField "IO Field_98" at 816,197 size 112x38; FormatPattern 99.99
      ProcessValue <- "ST_Calculation_Var_1_ZhiShu_ARRAY_JR{36}"
   IOField "IO Field_99" at 816,242 size 112x38; FormatPattern 99.99
      ProcessValue <- "ST_Calculation_Var_1_ZhiShu_ARRAY_JR{37}"
   IOField "IO Field_100" at 816,286 size 112x38; FormatPattern 99.99
      ProcessValue <- "ST_Calculation_Var_1_ZhiShu_ARRAY_JR{38}"
   IOField "IO Field_101" at 816,331 size 112x38; FormatPattern 99.99
      ProcessValue <- "ST_Calculation_Var_1_ZhiShu_ARRAY_JR{39}"
   IOField "IO Field_102" at 816,376 size 112x38; FormatPattern 99.99
      ProcessValue <- "ST_Calculation_Var_1_ZhiShu_ARRAY_JR{40}"
   IOField "IO Field_103" at 816,420 size 112x38; FormatPattern 99.99
      ProcessValue <- "ST_Calculation_Var_1_ZhiShu_ARRAY_JR{41}"
   IOField "IO Field_104" at 816,465 size 112x38; FormatPattern 99.99
      ProcessValue <- "ST_Calculation_Var_1_ZhiShu_ARRAY_JR{42}"
   IOField "IO Field_105" at 816,509 size 112x38; FormatPattern 99.99
      ProcessValue <- "ST_Calculation_Var_1_ZhiShu_ARRAY_JR{43}"
   IOField "IO Field_106" at 816,554 size 112x38; FormatPattern 99.99
      ProcessValue <- "ST_Calculation_Var_1_ZhiShu_ARRAY_JR{44}"
   IOField "IO Field_107" at 816,598 size 112x38; FormatPattern 99.99
      ProcessValue <- "ST_Calculation_Var_1_ZhiShu_ARRAY_JR{45}"
   IOField "IO Field_108" at 816,643 size 112x38; FormatPattern 99.99
      ProcessValue <- "ST_Calculation_Var_1_ZhiShu_ARRAY_JR{46}"
   IOField "IO Field_109" at 816,688 size 112x38; FormatPattern 99.99
      ProcessValue <- "ST_Calculation_Var_1_ZhiShu_ARRAY_JR{47}"
   IOField "IO Field_110" at 948,153 size 112x38; FormatPattern 99.999
      ProcessValue <- "ST_Calculation_Var_1_f1_n_delt_0_n_ARRAY_JR{35}"
   IOField "IO Field_111" at 948,197 size 112x38; FormatPattern 99.999
      ProcessValue <- "ST_Calculation_Var_1_f1_n_delt_0_n_ARRAY_JR{36}"
   IOField "IO Field_112" at 948,242 size 112x38; FormatPattern 99.999
      ProcessValue <- "ST_Calculation_Var_1_f1_n_delt_0_n_ARRAY_JR{37}"
   IOField "IO Field_113" at 948,286 size 112x38; FormatPattern 99.999
      ProcessValue <- "ST_Calculation_Var_1_f1_n_delt_0_n_ARRAY_JR{38}"
   IOField "IO Field_114" at 948,331 size 112x38; FormatPattern 99.999
      ProcessValue <- "ST_Calculation_Var_1_f1_n_delt_0_n_ARRAY_JR{39}"
   IOField "IO Field_115" at 948,376 size 112x38; FormatPattern 99.999
      ProcessValue <- "ST_Calculation_Var_1_f1_n_delt_0_n_ARRAY_JR{40}"
   IOField "IO Field_116" at 948,420 size 112x38; FormatPattern 99.999
      ProcessValue <- "ST_Calculation_Var_1_f1_n_delt_0_n_ARRAY_JR{41}"
   IOField "IO Field_117" at 948,465 size 112x38; FormatPattern 99.999
      ProcessValue <- "ST_Calculation_Var_1_f1_n_delt_0_n_ARRAY_JR{42}"
   IOField "IO Field_118" at 948,509 size 112x38; FormatPattern 99.999
      ProcessValue <- "ST_Calculation_Var_1_f1_n_delt_0_n_ARRAY_JR{43}"
   IOField "IO Field_119" at 948,554 size 112x38; FormatPattern 99.999
      ProcessValue <- "ST_Calculation_Var_1_f1_n_delt_0_n_ARRAY_JR{44}"
   IOField "IO Field_120" at 948,598 size 112x38; FormatPattern 99.999
      ProcessValue <- "ST_Calculation_Var_1_f1_n_delt_0_n_ARRAY_JR{45}"
   IOField "IO Field_121" at 948,643 size 112x38; FormatPattern 99.999
      ProcessValue <- "ST_Calculation_Var_1_f1_n_delt_0_n_ARRAY_JR{46}"
   IOField "IO Field_122" at 948,688 size 112x38; FormatPattern 99.999
      ProcessValue <- "ST_Calculation_Var_1_f1_n_delt_0_n_ARRAY_JR{47}"
   IOField "IO Field_123" at 1080,153 size 112x38; FormatPattern 99.999
      ProcessValue <- "ST_Calculation_Var_1_g1_n_delt_0_n_ARRAY_JR{35}"
   IOField "IO Field_124" at 1080,197 size 112x38; FormatPattern 99.999
      ProcessValue <- "ST_Calculation_Var_1_g1_n_delt_0_n_ARRAY_JR{36}"
   IOField "IO Field_125" at 1080,242 size 112x38; FormatPattern 99.999
      ProcessValue <- "ST_Calculation_Var_1_g1_n_delt_0_n_ARRAY_JR{37}"
   IOField "IO Field_126" at 1080,286 size 112x38; FormatPattern 99.999
      ProcessValue <- "ST_Calculation_Var_1_g1_n_delt_0_n_ARRAY_JR{38}"
   IOField "IO Field_127" at 1080,331 size 112x38; FormatPattern 99.999
      ProcessValue <- "ST_Calculation_Var_1_g1_n_delt_0_n_ARRAY_JR{39}"
   IOField "IO Field_128" at 1080,376 size 112x38; FormatPattern 99.999
      ProcessValue <- "ST_Calculation_Var_1_g1_n_delt_0_n_ARRAY_JR{40}"
   IOField "IO Field_129" at 1080,420 size 112x38; FormatPattern 99.999
      ProcessValue <- "ST_Calculation_Var_1_g1_n_delt_0_n_ARRAY_JR{41}"
   IOField "IO Field_130" at 1080,465 size 112x38; FormatPattern 99.999
      ProcessValue <- "ST_Calculation_Var_1_g1_n_delt_0_n_ARRAY_JR{42}"
   IOField "IO Field_131" at 1080,509 size 112x38; FormatPattern 99.999
      ProcessValue <- "ST_Calculation_Var_1_g1_n_delt_0_n_ARRAY_JR{43}"
   IOField "IO Field_132" at 1080,554 size 112x38; FormatPattern 99.999
      ProcessValue <- "ST_Calculation_Var_1_g1_n_delt_0_n_ARRAY_JR{44}"
   IOField "IO Field_133" at 1080,598 size 112x38; FormatPattern 99.999
      ProcessValue <- "ST_Calculation_Var_1_g1_n_delt_0_n_ARRAY_JR{45}"
   IOField "IO Field_134" at 1080,643 size 112x38; FormatPattern 99.999
      ProcessValue <- "ST_Calculation_Var_1_g1_n_delt_0_n_ARRAY_JR{46}"
   IOField "IO Field_135" at 1084,688 size 112x38; FormatPattern 99.999
      ProcessValue <- "ST_Calculation_Var_1_g1_n_delt_0_n_ARRAY_JR{47}"
   Button "OBJECT_3" at 24,8 size 112x48; TextOff '支数: / EXIT / 標準糸管１: / 표준보빈1:'
      on Press: SetTag("ST_HMI_Var_HMI_i16_Status_ShaGuan_Select", 1)
      Appearance <- "ST_HMI_Var_HMI_i16_Status_ShaGuan_Select"
   Button "OBJECT_1" at 156,8 size 112x48; TextOff 'f1_n: / EXIT / 標準糸管１: / 표준보빈1:'
      on Press: SetTag("ST_HMI_Var_HMI_i16_Status_ShaGuan_Select", 1)
      Appearance <- "ST_HMI_Var_HMI_i16_Status_ShaGuan_Select"
   Button "OBJECT_2" at 288,8 size 112x48; TextOff 'g1_n: / EXIT / 標準糸管１: / 표준보빈1:'
      on Press: SetTag("ST_HMI_Var_HMI_i16_Status_ShaGuan_Select", 1)
      Appearance <- "ST_HMI_Var_HMI_i16_Status_ShaGuan_Select"
   Button "OBJECT_4" at 420,8 size 112x48; TextOff '支数: / EXIT / 標準糸管１: / 표준보빈1:'
      on Press: SetTag("ST_HMI_Var_HMI_i16_Status_ShaGuan_Select", 1)
      Appearance <- "ST_HMI_Var_HMI_i16_Status_ShaGuan_Select"
   Button "OBJECT_5" at 552,8 size 112x48; TextOff 'f1_n: / EXIT / 標準糸管１: / 표준보빈1:'
      on Press: SetTag("ST_HMI_Var_HMI_i16_Status_ShaGuan_Select", 1)
      Appearance <- "ST_HMI_Var_HMI_i16_Status_ShaGuan_Select"
   Button "OBJECT_6" at 684,8 size 112x48; TextOff 'g1_n: / EXIT / 標準糸管１: / 표준보빈1:'
      on Press: SetTag("ST_HMI_Var_HMI_i16_Status_ShaGuan_Select", 1)
      Appearance <- "ST_HMI_Var_HMI_i16_Status_ShaGuan_Select"
   Button "OBJECT_7" at 816,8 size 112x48; TextOff '支数: / EXIT / 標準糸管１: / 표준보빈1:'
      on Press: SetTag("ST_HMI_Var_HMI_i16_Status_ShaGuan_Select", 1)
      Appearance <- "ST_HMI_Var_HMI_i16_Status_ShaGuan_Select"
   Button "OBJECT_8" at 948,8 size 112x48; TextOff 'f1_n: / EXIT / 標準糸管１: / 표준보빈1:'
      on Press: SetTag("ST_HMI_Var_HMI_i16_Status_ShaGuan_Select", 1)
      Appearance <- "ST_HMI_Var_HMI_i16_Status_ShaGuan_Select"
   Button "OBJECT_9" at 1080,8 size 112x48; TextOff 'g1_n: / EXIT / 標準糸管１: / 표준보빈1:'
      on Press: SetTag("ST_HMI_Var_HMI_i16_Status_ShaGuan_Select", 1)
      Appearance <- "ST_HMI_Var_HMI_i16_Status_ShaGuan_Select"

screen "生头相关" 1280x733, template "模板_2"
   on GenerateScreen: "TitleUpdater"()
   Button "HmiScreenItemData_1" at 1119,8 size 159x47; TextOn '向后'; TextOff '向后'
      on Release: ActivateScreen("常用调试画面", 0)
   TextField "Text Field_8" at 162,16 size 332x42; Text '1.毛轴头数'
   TextField "Text Field_9" at 162,72 size 332x42; Text '2.成形弓上升量'
   TextField "Text Field_10" at 408,424 size 264x42; Text '7.走车第一次回车量'
   TextField "Text Field_11" at 408,480 size 264x42; Text '8.纱管底部纱线卷绕长度'
   TextField "Text Field_12" at 408,536 size 264x42; Text '9.锭子走车传动比'
   TextField "Text Field_16" at 162,128 size 332x42; Text '3.回绕出车展距'
   TextField "Text Field_17" at 162,184 size 332x42; Text '4.回绕牵伸'
   TextField "Text Field_18" at 162,240 size 332x42; Text '5.回绕锭子走车传动比'
   TextField "Text Field_1" at 162,296 size 332x42; Text '6.生头起点位置'
   TextField "Text Field_2" at 24,384 size 112x32; Text '空锭(先插管)'
   TextField "Text Field_3" at 152,384 size 112x32; Text '空锭(光锭)'
   TextField "Text Field_4" at 280,384 size 112x32; Text '落纱生头'
   IOField "IO Field_41" at 24,16 size 112x42; FormatPattern 99
      ProcessValue <- "ST_HMI_Var_HMI_r64_MaoZhou_TouShu"
   IOField "IO Field_46" at 24,424 size 112x42; FormatPattern 999
      ProcessValue <- "ST_HMI_Var_HMI_r64Axis_ZouChe_Position_KongDing_8"
   IOField "IO Field_1" at 24,72 size 112x42; FormatPattern 99
      ProcessValue <- "ST_HMI_Var_HMI_r64Axis_ChengXing_Position_delt_KongDing_8"
   IOField "IO Field_2" at 24,536 size 112x42; FormatPattern 99.9
      ProcessValue <- "ST_HMI_Var_HMI_r64_DingZi_Zouche_ratio_KongDing_9"
   IOField "IO Field_3" at 280,424 size 112x42; FormatPattern 999
      ProcessValue <- "ST_HMI_Var_HMI_r64Axis_ZouChe_Position_LuoSha_8"
   IOField "IO Field_4" at 280,536 size 112x42; FormatPattern 99.9
      ProcessValue <- "ST_HMI_Var_HMI_r64_DingZi_Zouche_ratio_LuoSha_9"
   IOField "IO Field_6" at 24,480 size 112x42; FormatPattern 999
      ProcessValue <- "ST_HMI_Var_HMI_r64Axis_ZouChe_Position_KongDing_9"
   IOField "IO Field_5" at 216,480 size 112x42; FormatPattern 999
      ProcessValue <- "ST_HMI_Var_HMI_r64Axis_ZouChe_Position_LuoSha_9"
   IOField "IO Field_7" at 24,128 size 112x42; FormatPattern 999.9
      ProcessValue <- "ST_HMI_Var_HMI_r64Position_ChuChe_KongDing_65"
   IOField "IO Field_8" at 24,184 size 112x42; FormatPattern 9.99
      ProcessValue <- "ST_HMI_Var_HMI_r64QianShen_KongDing_65"
   IOField "IO Field_9" at 24,240 size 112x42; FormatPattern 99.9
      ProcessValue <- "ST_HMI_Var_HMI_r64_DingZi_Zouche_ratio_KongDing_65"
   IOField "IO Field_10" at 24,296 size 112x42; FormatPattern 99.9
      ProcessValue <- "ST_HMI_Var_HMI_r64Axis_ZouChe_Position_ShengTou_Start_Position"
   IOField "IO Field_11" at 152,424 size 112x42; FormatPattern 999
      ProcessValue <- "ST_HMI_Var_HMI_r64Axis_ZouChe_Position_KongDing_8_1"
   IOField "IO Field_12" at 152,536 size 112x42; FormatPattern 99.9
      ProcessValue <- "ST_HMI_Var_HMI_r64_DingZi_Zouche_ratio_KongDing_9_1"

VB script "Shasui"
   '注意：要启动脚本，请按下 <Ctrl><空格>，然后就可以看到各种不同函数。
   '通过使用系统函数或 WinCC flexible 对象模型来编写脚本。您可以通过 HMI 运行系统对象很容易地访问系统
   '。挑选对象引用的一个很便利的
   '方式是按下 <Alt><右箭头>。通过使用编程语言 VBScript 的基本功能部件
   '来设计复杂的脚本，并可以直接通过名称，例如 tag = 5，来访问变量。
   
   Dim a
   a=CDbl(SmartTags("ST_Main_Var_g_u16_N_Cycle_Single(1)")) 
   If a<= SmartTags("ST_FC_Var_g_ND") Then 
   	SmartTags("VBS_hengsi_status0")=Int(a/SmartTags("ST_FC_Var_g_ND")*25)
   	SmartTags("VBS_hengsi_status1")=80
   Else
   	SmartTags("VBS_hengsi_status1")=Int((a-SmartTags("ST_FC_Var_g_ND"))/(SmartTags("ST_FC_Var_g_N")-SmartTags("ST_FC_Var_g_ND"))*43)
   	SmartTags("VBS_hengsi_status0")=30
   	
   End If
   
   If SmartTags("ST_Main_Var_g_i16_Mode_Enabled")=512  Then 
   	SmartTags("VBS_hengsi_status1")=80
   	SmartTags("VBS_hengsi_status0")=30
   End If

VB script "timeConverse"
   '注意：要启动脚本，请按下 <Ctrl><空格>，然后就可以看到各种不同函数。
   '通过使用系统函数或 WinCC flexible 对象模型来编写脚本。您可以通过 HMI 运行系统对象很容易地访问系统
   '。挑选对象引用的一个很便利的
   '方式是按下 <Alt><右箭头>。通过使用编程语言 VBScript 的基本功能部件
   '来设计复杂的脚本，并可以直接通过名称，例如 tag = 5，来访问变量。
   'SmartTags("VBS_time_all_hour") = SmartTags("D435_ST_Maintenance_g_r64_Time_All")/3600 
   
   Dim a,b,c,d,e,f
   
   a = SmartTags("ST_Maintenance_g_r64_Time_All")/31536000
   SmartTags("VBS_time_year")=Int(a)
   
   
   b = (a - Int(a))*365
   SmartTags("VBS_time_day")=Int(b)
   
   c =( b - Int(b))*24 
   SmartTags("VBS_time_hour")=Int(c) 
   
   d = (c - Int(c))*60
   SmartTags("VBS_time_min")=Int(d)
   
   e = (d - Int(d))*60
   SmartTags("VBS_time_sec") = Int(e)
    
      
   'SmartTags("VBS_date1") = DateDiff("s", SmartTags("D435_ST_Main_Var_g_dateAndTime0"),Now)
   'SmartTags("VBS_runningRate")= SmartTags("D435_ST_Maintenance_g_r64_Time_All")  / SmartTags("VBS_date1") *100

VB script "TitleUpdater"
   Dim title
   Set title = HmiRuntime.Screens(0).ScreenItems("画面标题")
   title.Text = HmiRuntime.BaseScreenName

scheduled task "Job_1"
   on Action: function_f41c6f6c("user_name")

scheduled task "作业_3"
   on Action: ResetBit("VBS_alwaysFalse")
   Triggers <- "1 h"

scheduled task "Task_1"
   on Action: "Shasui"()
   Triggers <- "1 min"

scheduled task "Task_2"
   on Action: "timeConverse"()
*)

(* ===== HMI "HMI_RT_1" =====

ScreenModuleEditorView "面板_1(2)" 640x480
   Group "Group" at 10,10 size 111x159
*)

(* ===== HMI "WinCC flexible RT" =====
system functions are stored by id; their names below are inferred from use
connection "HMI_连接_1": ETHERNET, SIMOTION

